(* Logix 5000 project; controller MV vendor 1 type 14 code 217 rev 31.11; software revision 31.00; part 15 of 53 *)
(* tags used below, declared in another part *)
   CWD : CHECKWORD_FLAGS;
   MC_Delphi_I : DINT[60];
   MC_LTX_001_1 : PlantItem;   // LTX_001_1
   MC_LTX_001_1_RawInput : ALIAS FOR RIO_Rack_2:12:I.Data.16;   // MC_LTX_001_1
   MC_LTX_001_2 : PlantItem;   // LTX_001_2
   MC_LTX_001_2_RawInput : ALIAS FOR RIO_Rack_2:12:I.Data.17;   // MC_LTX_001_2
   MC_LTX_001_3 : PlantItem;   // LTX_001_3
   MC_LTX_001_3_RawInput : ALIAS FOR RIO_Rack_2:12:I.Data.18;   // MC_LTX_001_3
   MC_LTX_002_1 : PlantItem;   // LTX_002_1
   MC_LTX_002_1_RawInput : ALIAS FOR RIO_Rack_2:12:I.Data.19;   // MC_LTX_002_1
   MC_LTX_002_2 : PlantItem;   // LTX_002_2
   MC_LTX_002_2_RawInput : ALIAS FOR RIO_Rack_2:12:I.Data.20;   // MC_LTX_002_2
   MC_LTX_002_3 : PlantItem;   // LTX_002_3
   MC_LTX_002_3_RawInput : ALIAS FOR RIO_Rack_2:12:I.Data.21;   // MC_LTX_002_3
   MC_LTX_003_1 : PlantItem;   // LTX_003_1
   MC_LTX_003_1_RawInput : ALIAS FOR RIO_Rack_2:12:I.Data.22;   // MC_LTX_003_1
   MC_LTX_003_2 : PlantItem;   // LTX_003_2
   MC_LTX_003_2_RawInput : ALIAS FOR RIO_Rack_2:12:I.Data.23;   // MC_LTX_003_2
   MC_LTX_003_3 : PlantItem;   // LTX_003_3
   MC_LTX_003_3_RawInput : ALIAS FOR RIO_Rack_2:12:I.Data.24;   // MC_LTX_003_3
   MC_PILZ : PlantItem;   // PILZ
   MC_PILZ_RawInput : ALIAS FOR RIO_Rack_2:12:I.Data.31;   // MC_PILZ
   MC_PROXY2 : PlantItem;   // PROXY2
   MC_PROXY2_RawInput : ALIAS FOR RIO_Rack_2:12:I.Data.30;   // MC_PROXY2
   MC_PROXY_RawInput : ALIAS FOR RIO_Rack_2:12:I.Data.14;   // MC_PROXY
   MC_R3_SW2_1 : PlantItem;   // PROXY
   MC_R3_SW3 : PlantItem;   // R3_SW3
   MC_R3_SW3_RawInput : ALIAS FOR RIO_Rack_2:12:I.Data.7;   // MC_R3_SW3
   MC_R4_SW1 : PlantItem;   // R4_SW1
   MC_R4_SW1_RawInput : ALIAS FOR RIO_Rack_2:12:I.Data.8;   // MC_R4_SW1
   MC_R4_SW2 : PlantItem;   // R4_SW2
   MC_R4_SW2_RawInput : ALIAS FOR RIO_Rack_2:12:I.Data.9;   // MC_R4_SW2
   MC_R4_SW3 : PlantItem;   // R4_SW3
   MC_R4_SW3_RawInput : ALIAS FOR RIO_Rack_2:12:I.Data.10;   // MC_R4_SW3
   MC_R4_SW4 : PlantItem;   // R4_SW4
   MC_R4_SW4_RawInput : ALIAS FOR RIO_Rack_2:12:I.Data.11;   // MC_R4_SW4
   MC_R4_SW6 : PlantItem;   // R4_SW6
   MC_R4_SW6_RawInput : ALIAS FOR RIO_Rack_2:12:I.Data.12;   // MC_R4_SW6
   MC_R6_SW1 : PlantItem;   // R6_SW1
   MC_R6_SW1_RawInput : ALIAS FOR RIO_Rack_2:12:I.Data.13;   // MC_R6_SW1
   One_Second_One_Scan : ALIAS FOR One_Second_1_scan;
(* MC_Common, continued *)

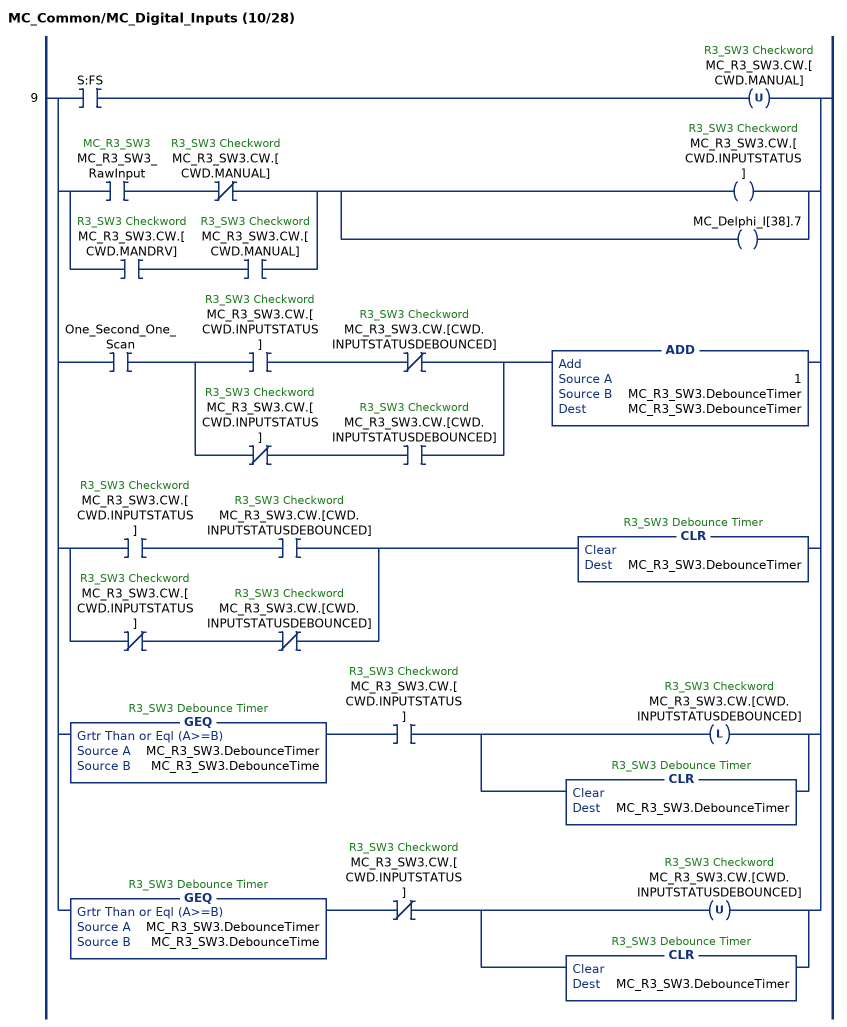
   [picture p227: MC_Common/MC_Digital_Inputs rungs 9-9]
   9: [XIC(S:FS) OTU(MC_R3_SW3.CW.[CWD.MANUAL]) ,[XIC(MC_R3_SW3_RawInput) XIO(MC_R3_SW3.CW.[CWD.MANUAL]) ,XIC(MC_R3_SW3.CW.[CWD.MANDRV]) XIC(MC_R3_SW3.CW.[CWD.MANUAL]) ] [OTE(MC_R3_SW3.CW.[CWD.INPUTSTATUS]) ,OTE(MC_Delphi_I[38].7) ] ,XIC(One_Second_One_Scan) [XIC(MC_R3_SW3.CW.[CWD.INPUTSTATUS]) XIO(MC_R3_SW3.CW.[CWD.INPUTSTATUSDEBOUNCED]) ,XIO(MC_R3_SW3.CW.[CWD.INPUTSTATUS]) XIC(MC_R3_SW3.CW.[CWD.INPUTSTATUSDEBOUNCED]) ] ADD(1,MC_R3_SW3.DebounceTimer,MC_R3_SW3.DebounceTimer) ,[XIC(MC_R3_SW3.CW.[CWD.INPUTSTATUS]) XIC(MC_R3_SW3.CW.[CWD.INPUTSTATUSDEBOUNCED]) ,XIO(MC_R3_SW3.CW.[CWD.INPUTSTATUS]) XIO(MC_R3_SW3.CW.[CWD.INPUTSTATUSDEBOUNCED]) ] CLR(MC_R3_SW3.DebounceTimer) ,GEQ(MC_R3_SW3.DebounceTimer,MC_R3_SW3.DebounceTime) XIC(MC_R3_SW3.CW.[CWD.INPUTSTATUS]) [OTL(MC_R3_SW3.CW.[CWD.INPUTSTATUSDEBOUNCED]) ,CLR(MC_R3_SW3.DebounceTimer) ] ,GEQ(MC_R3_SW3.DebounceTimer,MC_R3_SW3.DebounceTime) XIO(MC_R3_SW3.CW.[CWD.INPUTSTATUS]) [OTU(MC_R3_SW3.CW.[CWD.INPUTSTATUSDEBOUNCED]) ,CLR(MC_R3_SW3.DebounceTimer) ] ];
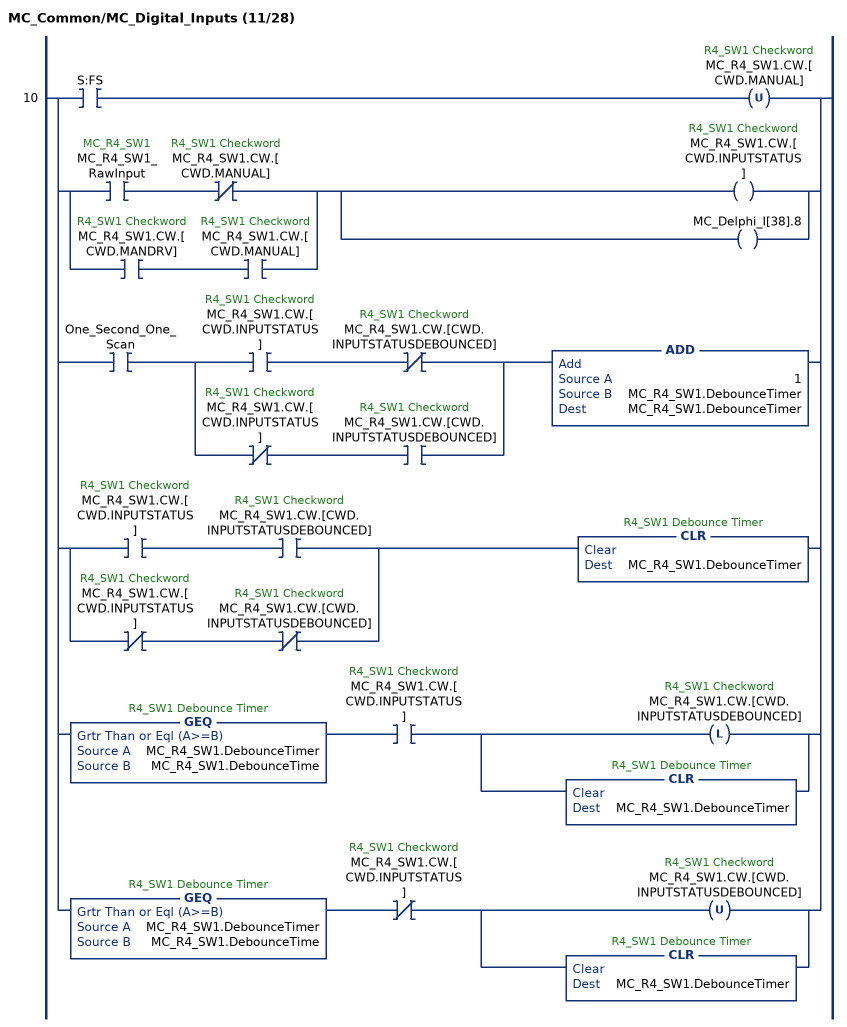
   10: [XIC(S:FS) OTU(MC_R4_SW1.CW.[CWD.MANUAL]) ,[XIC(MC_R4_SW1_RawInput) XIO(MC_R4_SW1.CW.[CWD.MANUAL]) ,XIC(MC_R4_SW1.CW.[CWD.MANDRV]) XIC(MC_R4_SW1.CW.[CWD.MANUAL]) ] [OTE(MC_R4_SW1.CW.[CWD.INPUTSTATUS]) ,OTE(MC_Delphi_I[38].8) ] ,XIC(One_Second_One_Scan) [XIC(MC_R4_SW1.CW.[CWD.INPUTSTATUS]) XIO(MC_R4_SW1.CW.[CWD.INPUTSTATUSDEBOUNCED]) ,XIO(MC_R4_SW1.CW.[CWD.INPUTSTATUS]) XIC(MC_R4_SW1.CW.[CWD.INPUTSTATUSDEBOUNCED]) ] ADD(1,MC_R4_SW1.DebounceTimer,MC_R4_SW1.DebounceTimer) ,[XIC(MC_R4_SW1.CW.[CWD.INPUTSTATUS]) XIC(MC_R4_SW1.CW.[CWD.INPUTSTATUSDEBOUNCED]) ,XIO(MC_R4_SW1.CW.[CWD.INPUTSTATUS]) XIO(MC_R4_SW1.CW.[CWD.INPUTSTATUSDEBOUNCED]) ] CLR(MC_R4_SW1.DebounceTimer) ,GEQ(MC_R4_SW1.DebounceTimer,MC_R4_SW1.DebounceTime) XIC(MC_R4_SW1.CW.[CWD.INPUTSTATUS]) [OTL(MC_R4_SW1.CW.[CWD.INPUTSTATUSDEBOUNCED]) ,CLR(MC_R4_SW1.DebounceTimer) ] ,GEQ(MC_R4_SW1.DebounceTimer,MC_R4_SW1.DebounceTime) XIO(MC_R4_SW1.CW.[CWD.INPUTSTATUS]) [OTU(MC_R4_SW1.CW.[CWD.INPUTSTATUSDEBOUNCED]) ,CLR(MC_R4_SW1.DebounceTimer) ] ];
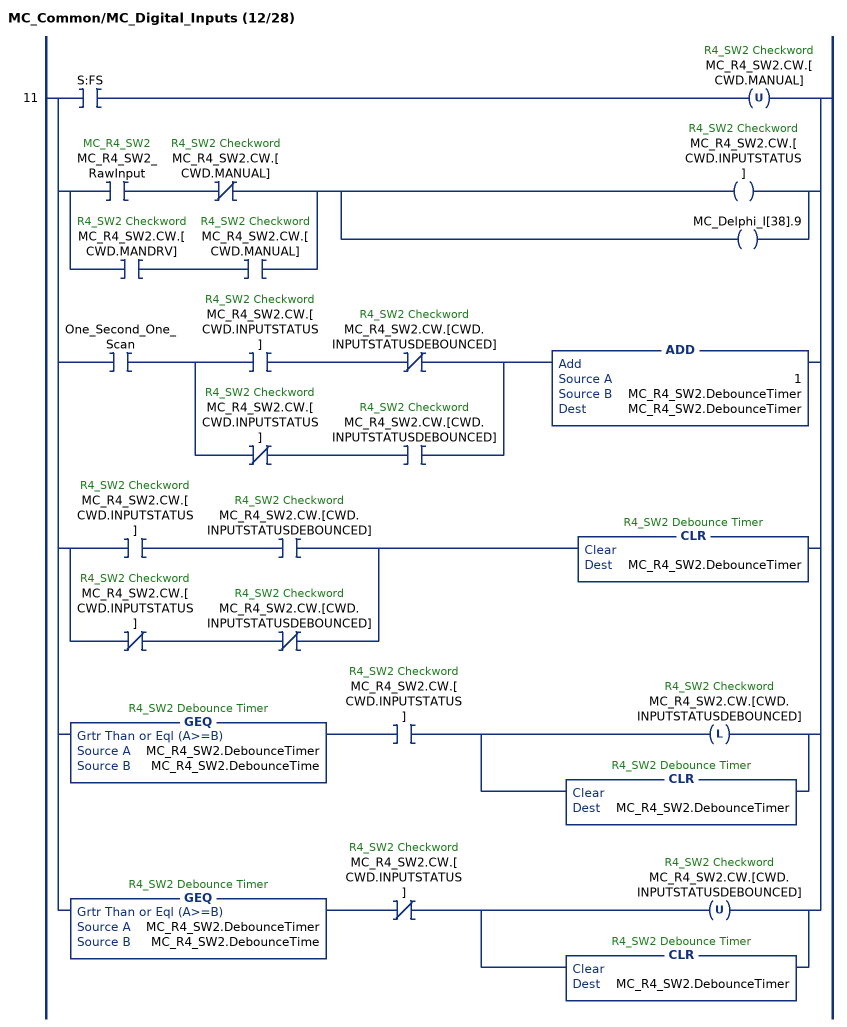
   11: [XIC(S:FS) OTU(MC_R4_SW2.CW.[CWD.MANUAL]) ,[XIC(MC_R4_SW2_RawInput) XIO(MC_R4_SW2.CW.[CWD.MANUAL]) ,XIC(MC_R4_SW2.CW.[CWD.MANDRV]) XIC(MC_R4_SW2.CW.[CWD.MANUAL]) ] [OTE(MC_R4_SW2.CW.[CWD.INPUTSTATUS]) ,OTE(MC_Delphi_I[38].9) ] ,XIC(One_Second_One_Scan) [XIC(MC_R4_SW2.CW.[CWD.INPUTSTATUS]) XIO(MC_R4_SW2.CW.[CWD.INPUTSTATUSDEBOUNCED]) ,XIO(MC_R4_SW2.CW.[CWD.INPUTSTATUS]) XIC(MC_R4_SW2.CW.[CWD.INPUTSTATUSDEBOUNCED]) ] ADD(1,MC_R4_SW2.DebounceTimer,MC_R4_SW2.DebounceTimer) ,[XIC(MC_R4_SW2.CW.[CWD.INPUTSTATUS]) XIC(MC_R4_SW2.CW.[CWD.INPUTSTATUSDEBOUNCED]) ,XIO(MC_R4_SW2.CW.[CWD.INPUTSTATUS]) XIO(MC_R4_SW2.CW.[CWD.INPUTSTATUSDEBOUNCED]) ] CLR(MC_R4_SW2.DebounceTimer) ,GEQ(MC_R4_SW2.DebounceTimer,MC_R4_SW2.DebounceTime) XIC(MC_R4_SW2.CW.[CWD.INPUTSTATUS]) [OTL(MC_R4_SW2.CW.[CWD.INPUTSTATUSDEBOUNCED]) ,CLR(MC_R4_SW2.DebounceTimer) ] ,GEQ(MC_R4_SW2.DebounceTimer,MC_R4_SW2.DebounceTime) XIO(MC_R4_SW2.CW.[CWD.INPUTSTATUS]) [OTU(MC_R4_SW2.CW.[CWD.INPUTSTATUSDEBOUNCED]) ,CLR(MC_R4_SW2.DebounceTimer) ] ];
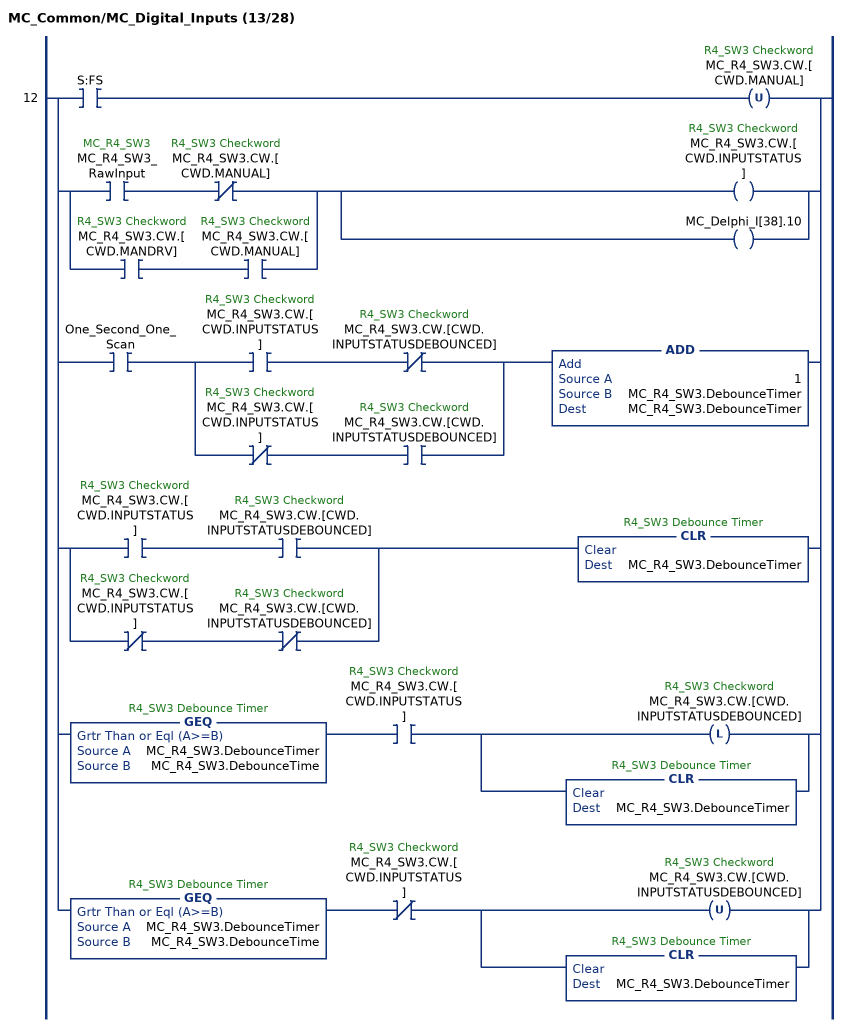
   12: [XIC(S:FS) OTU(MC_R4_SW3.CW.[CWD.MANUAL]) ,[XIC(MC_R4_SW3_RawInput) XIO(MC_R4_SW3.CW.[CWD.MANUAL]) ,XIC(MC_R4_SW3.CW.[CWD.MANDRV]) XIC(MC_R4_SW3.CW.[CWD.MANUAL]) ] [OTE(MC_R4_SW3.CW.[CWD.INPUTSTATUS]) ,OTE(MC_Delphi_I[38].10) ] ,XIC(One_Second_One_Scan) [XIC(MC_R4_SW3.CW.[CWD.INPUTSTATUS]) XIO(MC_R4_SW3.CW.[CWD.INPUTSTATUSDEBOUNCED]) ,XIO(MC_R4_SW3.CW.[CWD.INPUTSTATUS]) XIC(MC_R4_SW3.CW.[CWD.INPUTSTATUSDEBOUNCED]) ] ADD(1,MC_R4_SW3.DebounceTimer,MC_R4_SW3.DebounceTimer) ,[XIC(MC_R4_SW3.CW.[CWD.INPUTSTATUS]) XIC(MC_R4_SW3.CW.[CWD.INPUTSTATUSDEBOUNCED]) ,XIO(MC_R4_SW3.CW.[CWD.INPUTSTATUS]) XIO(MC_R4_SW3.CW.[CWD.INPUTSTATUSDEBOUNCED]) ] CLR(MC_R4_SW3.DebounceTimer) ,GEQ(MC_R4_SW3.DebounceTimer,MC_R4_SW3.DebounceTime) XIC(MC_R4_SW3.CW.[CWD.INPUTSTATUS]) [OTL(MC_R4_SW3.CW.[CWD.INPUTSTATUSDEBOUNCED]) ,CLR(MC_R4_SW3.DebounceTimer) ] ,GEQ(MC_R4_SW3.DebounceTimer,MC_R4_SW3.DebounceTime) XIO(MC_R4_SW3.CW.[CWD.INPUTSTATUS]) [OTU(MC_R4_SW3.CW.[CWD.INPUTSTATUSDEBOUNCED]) ,CLR(MC_R4_SW3.DebounceTimer) ] ];
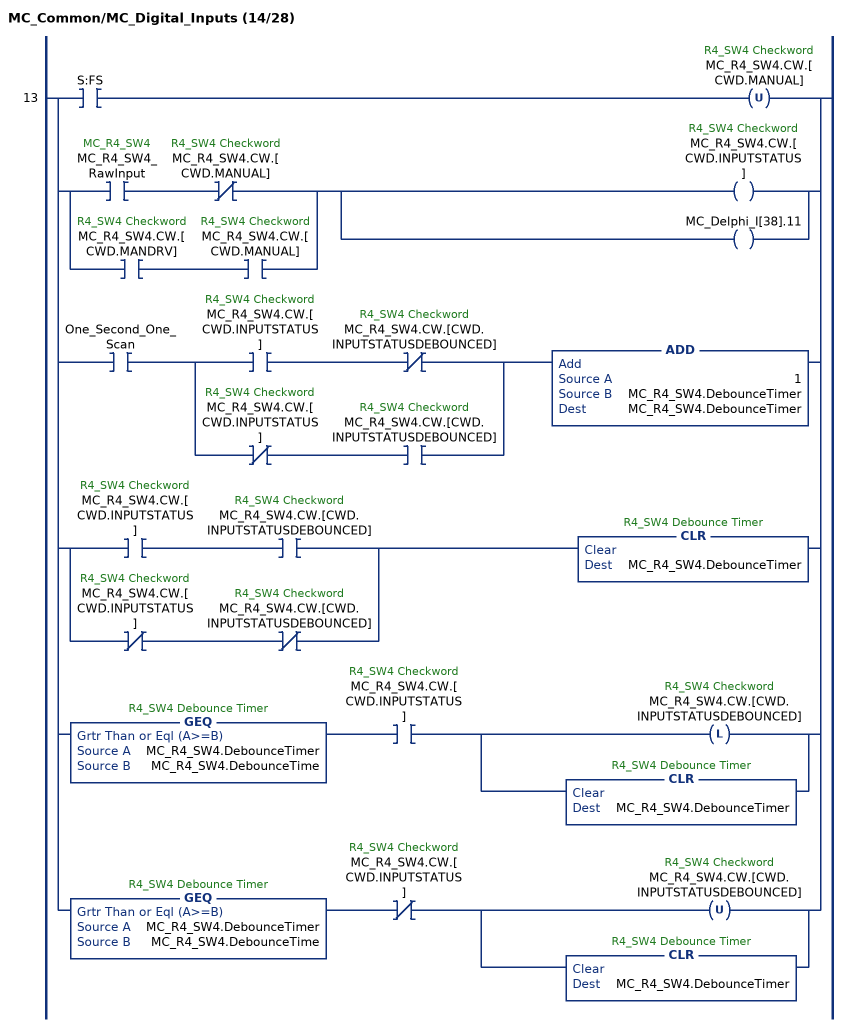
   13: [XIC(S:FS) OTU(MC_R4_SW4.CW.[CWD.MANUAL]) ,[XIC(MC_R4_SW4_RawInput) XIO(MC_R4_SW4.CW.[CWD.MANUAL]) ,XIC(MC_R4_SW4.CW.[CWD.MANDRV]) XIC(MC_R4_SW4.CW.[CWD.MANUAL]) ] [OTE(MC_R4_SW4.CW.[CWD.INPUTSTATUS]) ,OTE(MC_Delphi_I[38].11) ] ,XIC(One_Second_One_Scan) [XIC(MC_R4_SW4.CW.[CWD.INPUTSTATUS]) XIO(MC_R4_SW4.CW.[CWD.INPUTSTATUSDEBOUNCED]) ,XIO(MC_R4_SW4.CW.[CWD.INPUTSTATUS]) XIC(MC_R4_SW4.CW.[CWD.INPUTSTATUSDEBOUNCED]) ] ADD(1,MC_R4_SW4.DebounceTimer,MC_R4_SW4.DebounceTimer) ,[XIC(MC_R4_SW4.CW.[CWD.INPUTSTATUS]) XIC(MC_R4_SW4.CW.[CWD.INPUTSTATUSDEBOUNCED]) ,XIO(MC_R4_SW4.CW.[CWD.INPUTSTATUS]) XIO(MC_R4_SW4.CW.[CWD.INPUTSTATUSDEBOUNCED]) ] CLR(MC_R4_SW4.DebounceTimer) ,GEQ(MC_R4_SW4.DebounceTimer,MC_R4_SW4.DebounceTime) XIC(MC_R4_SW4.CW.[CWD.INPUTSTATUS]) [OTL(MC_R4_SW4.CW.[CWD.INPUTSTATUSDEBOUNCED]) ,CLR(MC_R4_SW4.DebounceTimer) ] ,GEQ(MC_R4_SW4.DebounceTimer,MC_R4_SW4.DebounceTime) XIO(MC_R4_SW4.CW.[CWD.INPUTSTATUS]) [OTU(MC_R4_SW4.CW.[CWD.INPUTSTATUSDEBOUNCED]) ,CLR(MC_R4_SW4.DebounceTimer) ] ];
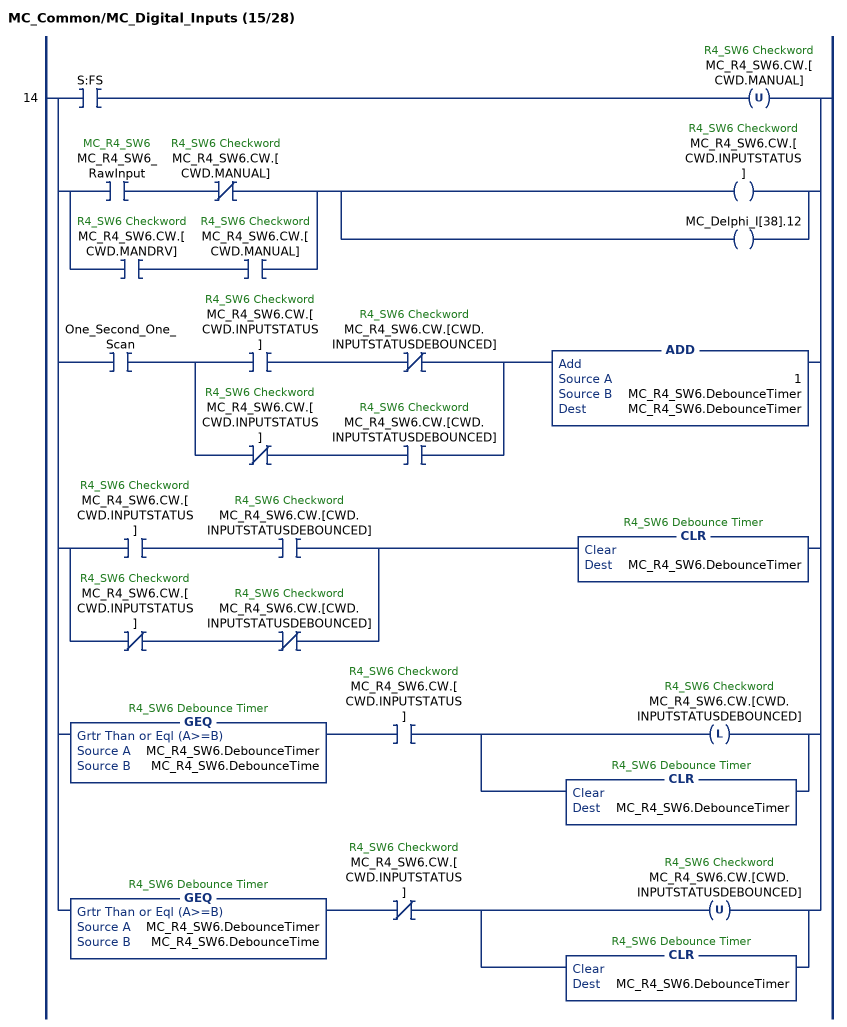
   14: [XIC(S:FS) OTU(MC_R4_SW6.CW.[CWD.MANUAL]) ,[XIC(MC_R4_SW6_RawInput) XIO(MC_R4_SW6.CW.[CWD.MANUAL]) ,XIC(MC_R4_SW6.CW.[CWD.MANDRV]) XIC(MC_R4_SW6.CW.[CWD.MANUAL]) ] [OTE(MC_R4_SW6.CW.[CWD.INPUTSTATUS]) ,OTE(MC_Delphi_I[38].12) ] ,XIC(One_Second_One_Scan) [XIC(MC_R4_SW6.CW.[CWD.INPUTSTATUS]) XIO(MC_R4_SW6.CW.[CWD.INPUTSTATUSDEBOUNCED]) ,XIO(MC_R4_SW6.CW.[CWD.INPUTSTATUS]) XIC(MC_R4_SW6.CW.[CWD.INPUTSTATUSDEBOUNCED]) ] ADD(1,MC_R4_SW6.DebounceTimer,MC_R4_SW6.DebounceTimer) ,[XIC(MC_R4_SW6.CW.[CWD.INPUTSTATUS]) XIC(MC_R4_SW6.CW.[CWD.INPUTSTATUSDEBOUNCED]) ,XIO(MC_R4_SW6.CW.[CWD.INPUTSTATUS]) XIO(MC_R4_SW6.CW.[CWD.INPUTSTATUSDEBOUNCED]) ] CLR(MC_R4_SW6.DebounceTimer) ,GEQ(MC_R4_SW6.DebounceTimer,MC_R4_SW6.DebounceTime) XIC(MC_R4_SW6.CW.[CWD.INPUTSTATUS]) [OTL(MC_R4_SW6.CW.[CWD.INPUTSTATUSDEBOUNCED]) ,CLR(MC_R4_SW6.DebounceTimer) ] ,GEQ(MC_R4_SW6.DebounceTimer,MC_R4_SW6.DebounceTime) XIO(MC_R4_SW6.CW.[CWD.INPUTSTATUS]) [OTU(MC_R4_SW6.CW.[CWD.INPUTSTATUSDEBOUNCED]) ,CLR(MC_R4_SW6.DebounceTimer) ] ];
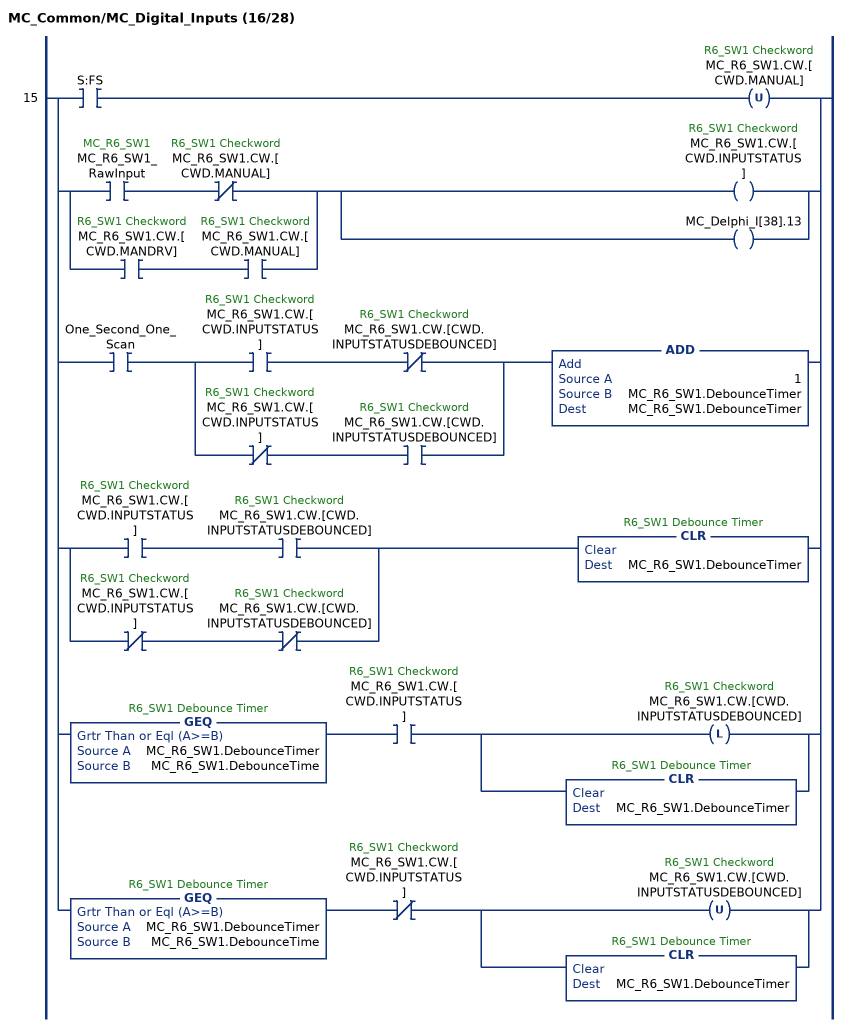
   15: [XIC(S:FS) OTU(MC_R6_SW1.CW.[CWD.MANUAL]) ,[XIC(MC_R6_SW1_RawInput) XIO(MC_R6_SW1.CW.[CWD.MANUAL]) ,XIC(MC_R6_SW1.CW.[CWD.MANDRV]) XIC(MC_R6_SW1.CW.[CWD.MANUAL]) ] [OTE(MC_R6_SW1.CW.[CWD.INPUTSTATUS]) ,OTE(MC_Delphi_I[38].13) ] ,XIC(One_Second_One_Scan) [XIC(MC_R6_SW1.CW.[CWD.INPUTSTATUS]) XIO(MC_R6_SW1.CW.[CWD.INPUTSTATUSDEBOUNCED]) ,XIO(MC_R6_SW1.CW.[CWD.INPUTSTATUS]) XIC(MC_R6_SW1.CW.[CWD.INPUTSTATUSDEBOUNCED]) ] ADD(1,MC_R6_SW1.DebounceTimer,MC_R6_SW1.DebounceTimer) ,[XIC(MC_R6_SW1.CW.[CWD.INPUTSTATUS]) XIC(MC_R6_SW1.CW.[CWD.INPUTSTATUSDEBOUNCED]) ,XIO(MC_R6_SW1.CW.[CWD.INPUTSTATUS]) XIO(MC_R6_SW1.CW.[CWD.INPUTSTATUSDEBOUNCED]) ] CLR(MC_R6_SW1.DebounceTimer) ,GEQ(MC_R6_SW1.DebounceTimer,MC_R6_SW1.DebounceTime) XIC(MC_R6_SW1.CW.[CWD.INPUTSTATUS]) [OTL(MC_R6_SW1.CW.[CWD.INPUTSTATUSDEBOUNCED]) ,CLR(MC_R6_SW1.DebounceTimer) ] ,GEQ(MC_R6_SW1.DebounceTimer,MC_R6_SW1.DebounceTime) XIO(MC_R6_SW1.CW.[CWD.INPUTSTATUS]) [OTU(MC_R6_SW1.CW.[CWD.INPUTSTATUSDEBOUNCED]) ,CLR(MC_R6_SW1.DebounceTimer) ] ];
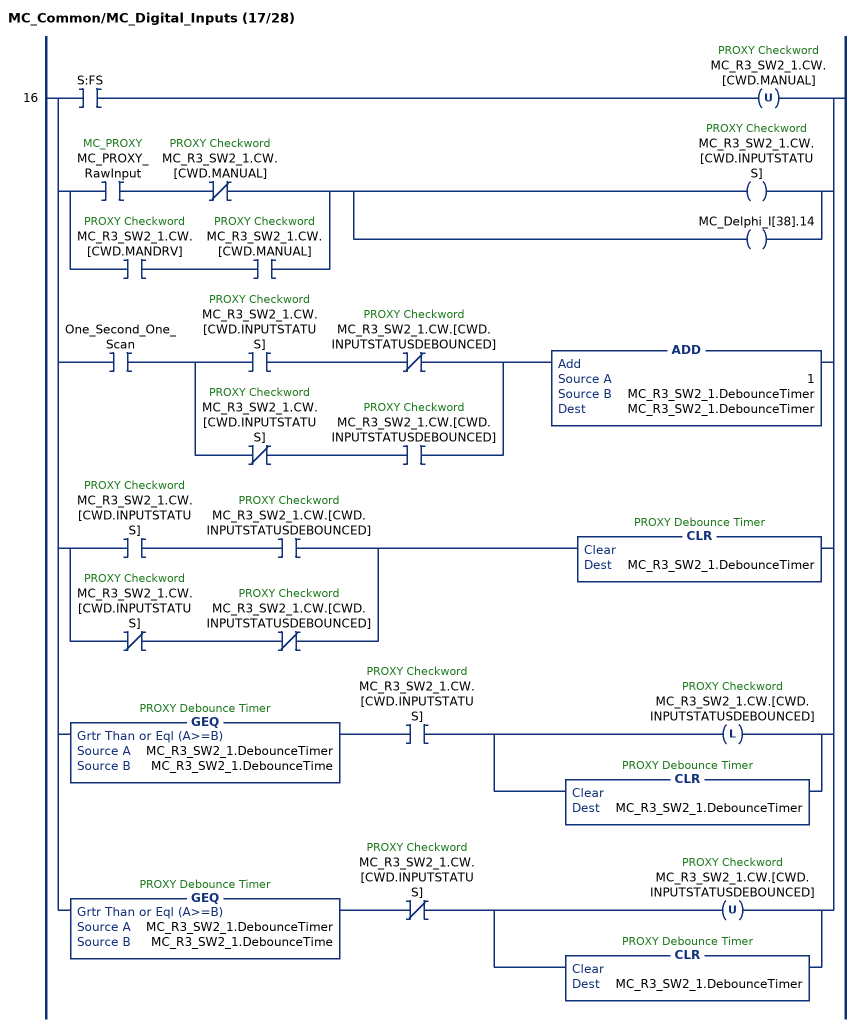
   16: [XIC(S:FS) OTU(MC_R3_SW2_1.CW.[CWD.MANUAL]) ,[XIC(MC_PROXY_RawInput) XIO(MC_R3_SW2_1.CW.[CWD.MANUAL]) ,XIC(MC_R3_SW2_1.CW.[CWD.MANDRV]) XIC(MC_R3_SW2_1.CW.[CWD.MANUAL]) ] [OTE(MC_R3_SW2_1.CW.[CWD.INPUTSTATUS]) ,OTE(MC_Delphi_I[38].14) ] ,XIC(One_Second_One_Scan) [XIC(MC_R3_SW2_1.CW.[CWD.INPUTSTATUS]) XIO(MC_R3_SW2_1.CW.[CWD.INPUTSTATUSDEBOUNCED]) ,XIO(MC_R3_SW2_1.CW.[CWD.INPUTSTATUS]) XIC(MC_R3_SW2_1.CW.[CWD.INPUTSTATUSDEBOUNCED]) ] ADD(1,MC_R3_SW2_1.DebounceTimer,MC_R3_SW2_1.DebounceTimer) ,[XIC(MC_R3_SW2_1.CW.[CWD.INPUTSTATUS]) XIC(MC_R3_SW2_1.CW.[CWD.INPUTSTATUSDEBOUNCED]) ,XIO(MC_R3_SW2_1.CW.[CWD.INPUTSTATUS]) XIO(MC_R3_SW2_1.CW.[CWD.INPUTSTATUSDEBOUNCED]) ] CLR(MC_R3_SW2_1.DebounceTimer) ,GEQ(MC_R3_SW2_1.DebounceTimer,MC_R3_SW2_1.DebounceTime) XIC(MC_R3_SW2_1.CW.[CWD.INPUTSTATUS]) [OTL(MC_R3_SW2_1.CW.[CWD.INPUTSTATUSDEBOUNCED]) ,CLR(MC_R3_SW2_1.DebounceTimer) ] ,GEQ(MC_R3_SW2_1.DebounceTimer,MC_R3_SW2_1.DebounceTime) XIO(MC_R3_SW2_1.CW.[CWD.INPUTSTATUS]) [OTU(MC_R3_SW2_1.CW.[CWD.INPUTSTATUSDEBOUNCED]) ,CLR(MC_R3_SW2_1.DebounceTimer) ] ];
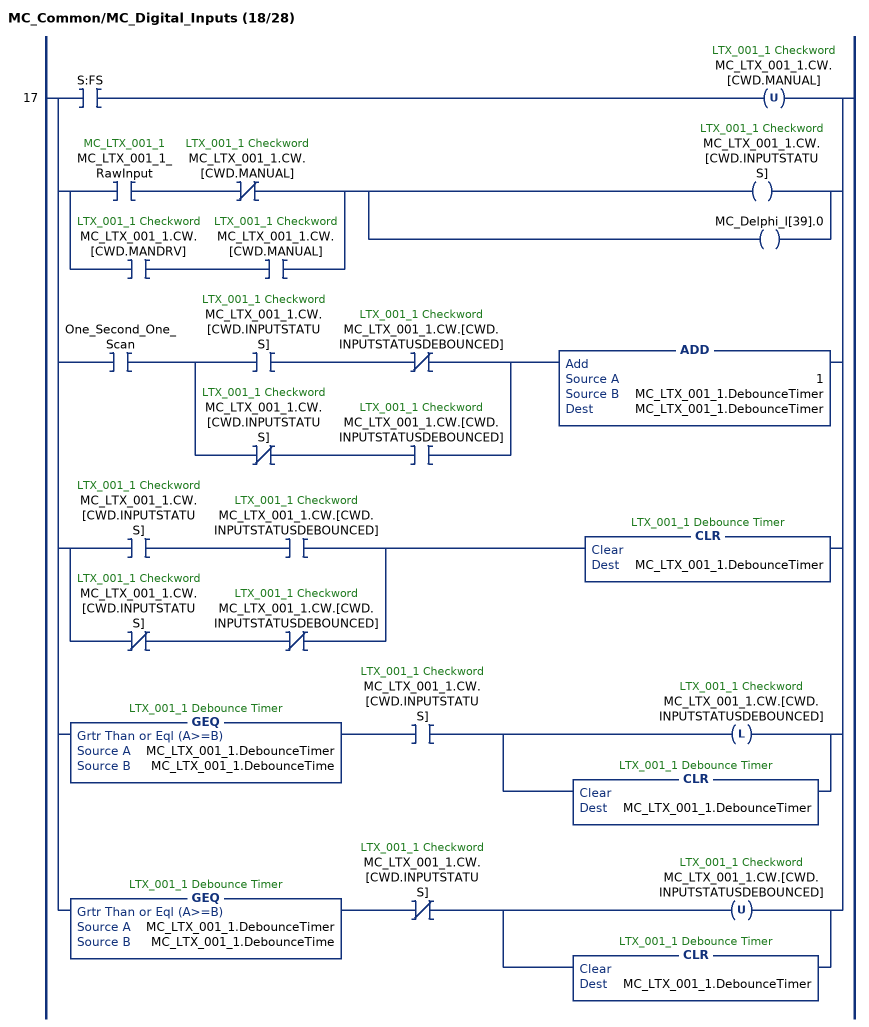
   17: [XIC(S:FS) OTU(MC_LTX_001_1.CW.[CWD.MANUAL]) ,[XIC(MC_LTX_001_1_RawInput) XIO(MC_LTX_001_1.CW.[CWD.MANUAL]) ,XIC(MC_LTX_001_1.CW.[CWD.MANDRV]) XIC(MC_LTX_001_1.CW.[CWD.MANUAL]) ] [OTE(MC_LTX_001_1.CW.[CWD.INPUTSTATUS]) ,OTE(MC_Delphi_I[39].0) ] ,XIC(One_Second_One_Scan) [XIC(MC_LTX_001_1.CW.[CWD.INPUTSTATUS]) XIO(MC_LTX_001_1.CW.[CWD.INPUTSTATUSDEBOUNCED]) ,XIO(MC_LTX_001_1.CW.[CWD.INPUTSTATUS]) XIC(MC_LTX_001_1.CW.[CWD.INPUTSTATUSDEBOUNCED]) ] ADD(1,MC_LTX_001_1.DebounceTimer,MC_LTX_001_1.DebounceTimer) ,[XIC(MC_LTX_001_1.CW.[CWD.INPUTSTATUS]) XIC(MC_LTX_001_1.CW.[CWD.INPUTSTATUSDEBOUNCED]) ,XIO(MC_LTX_001_1.CW.[CWD.INPUTSTATUS]) XIO(MC_LTX_001_1.CW.[CWD.INPUTSTATUSDEBOUNCED]) ] CLR(MC_LTX_001_1.DebounceTimer) ,GEQ(MC_LTX_001_1.DebounceTimer,MC_LTX_001_1.DebounceTime) XIC(MC_LTX_001_1.CW.[CWD.INPUTSTATUS]) [OTL(MC_LTX_001_1.CW.[CWD.INPUTSTATUSDEBOUNCED]) ,CLR(MC_LTX_001_1.DebounceTimer) ] ,GEQ(MC_LTX_001_1.DebounceTimer,MC_LTX_001_1.DebounceTime) XIO(MC_LTX_001_1.CW.[CWD.INPUTSTATUS]) [OTU(MC_LTX_001_1.CW.[CWD.INPUTSTATUSDEBOUNCED]) ,CLR(MC_LTX_001_1.DebounceTimer) ] ];